// TIA Portal project "OpenLibraryExample" (V13)

(* hardware
DEVICE "S71500/ET200MP station_1"  S7-1500 station
   slot 0: "Rail_0"  6ES7 590-1***0-0AA0
   slot 1: "WaterTreatmentPLC"  CPU 1516-3 PN/DP  6ES7 516-3AN01-0AB0  V1.8
   slot 2: "DI 16x24VDC BA_1"  DI 16x24VDC BA  6ES7 521-1BH10-0AA0  V1.0
   slot 3: "DQ 16x24VDC/0.5A BA_1"  DQ 16x24VDC/0.5A BA  6ES7 522-1BH10-0AA0  V1.0
   slot 4: "AI 4xU/I/RTD/TC ST_1"  AI 4xU/I/RTD/TC ST  6ES7 531-7QD00-0AB0  V1.0
   slot 5: "AQ 4xU/I ST_1"  AQ 4xU/I ST  6ES7 532-5HD00-0AB0  V2.0
DEVICE "SINAMICS G_1"  Sinamics.Device
   slot 0: "	_0"  Rail
   slot 0: "WaterPump"  G120 CU240E-2 PN  6SL3244-0BB12-1FA0  4.7.3
   slot 3: "PM240 IP20"  PM240 IP20  6SL3224-0BE31-5UA0  -
DEVICE "WaterTreatmentHMI"  TP900 Comfort
   slot 0: "HMI"  HMI  6AV2 124-0JC01-0AX0  13.0.1.0
   slot 1: "HMI_RT_1"  TP900 Comfort  6AV2 124-0JC01-0AX0  13.0.1.0
   slot 5: "WaterTreatmentHMI.IE_CP_1"  PROFINET Interface
      slot 1: "PROFINET Interface_1"  PROFINET Interface
         slot 1: "Port_1"  Port
         slot 2: "Port_2"  Port
   slot 7: "WaterTreatmentHMI.MPI/DP_CP_1"  MPI/DP Interface
*)

// ===== PLC "WaterTreatmentPLC"  CPU 1516-3 PN/DP =====

VAR_GLOBAL   // PLC tag table "Open Library"
   "System_Byte" AT %MB1 : Byte;
   "Clock_Byte" AT %MB0 : Byte;
   "Clock_10Hz" AT %M0.0 : Bool;
   "Clock_5Hz" AT %M0.1 : Bool;
   "Clock_2.5Hz" AT %M0.2 : Bool;
   "Clock_2Hz" AT %M0.3 : Bool;
   "Clock_1.25Hz" AT %M0.4 : Bool;
   "Clock_1Hz" AT %M0.5 : Bool;
   "Clock_0.625Hz" AT %M0.6 : Bool;
   "Clock_0.5Hz" AT %M0.7 : Bool;
   "AlwaysTRUE" AT %M1.2 : Bool;
   "AlwaysFALSE" AT %M1.3 : Bool;
   "FirstScan" AT %M1.0 : Bool;
   "DiagStatusUpdate" AT %M1.1 : Bool;
END_VAR

VAR_GLOBAL CONSTANT   // PLC tag table "Open Library"
   "Modes.Auto" : Int := 1;
   "Modes.Manual" : Int := 2;
   "Modes.Independent" : Int := 10;
   "Modes.Stop" : Int := 0;
   "HMI.Status.Stopped" : Int := 0;
   "HMI.Status.Estop" : Int := 1;
   "HMI.Status.Error" : Int := 2;
   "HMI.Status.ForwardWork" : Int := 3;
   "HMI.Status.ReverseHome" : Int := 4;
   "HMI.Status.OnForwardWork" : Int := 5;
   "HMI.Status.OnReverseHome" : Int := 6;
   "IoScaling.S7Analog.Default.iRawMax" : Int := 27648;
   "IoScaling.S7Analog.Default.iRawMin" : Int := 0;
   "IoScaling.S7Analog.Default.bSwapBytes" : Bool := false;
   "IoScaling.S7Analog.+-V/mA.iRawMax" : Int := 27648;
   "IoScaling.S7Analog.+-V/mA.iRawMin" : Int := -27648;
   "IoScaling.S7Analog.Types.Default" : Int := 0;
   "IoScaling.S7Analog.Pt100.iRawMax" : Int := 8500;
   "IoScaling.S7Analog.Pt100.iRawMin" : Int := -2000;
   "IoScaling.S7Analog.Pt100.Climate.iRawMax" : Int := 13000;
   "IoScaling.S7Analog.Pt100.Climate.iRawMin" : Int := -12000;
   "IoScaling.S7Analog.Ni100.iRawMax" : Int := 2500;
   "IoScaling.S7Analog.Ni100.iRawMin" : Int := -600;
   "IoScaling.S7Analog.Ni100.Climate.iRawMax" : Int := 25000;
   "IoScaling.S7Analog.Ni100.Climate.iRawMin" : Int := -6000;
   "IoScaling.S7Analog.Types.+-V/mA" : Int := 1;
   "IoScaling.S7Analog.Types.Pt100" : Int := 2;
   "IoScaling.S7Analog.Types.Pt100.Climate" : Int := 3;
   "IoScaling.S7Analog.Types.Ni100" : Int := 4;
   "IoScaling.S7Analog.Types.Ni100.Climate" : Int := 5;
   "IoScaling.S7Analog.Pt100.rScaledMax" : Real := 850.0;
   "IoScaling.S7Analog.Pt100.rScaledMin" : Real := -200.0;
   "IoScaling.S7Analog.Pt100.Climate.rScaledMax" : Real := 130.0;
   "IoScaling.S7Analog.Pt100.Climate.rScaledMin" : Real := -120.0;
   "IoScaling.S7Analog.Ni100.rScaledMax" : Real := 250.0;
   "IoScaling.S7Analog.Ni100.rScaledMin" : Real := -60.0;
   "IoScaling.S7Analog.Ni100.Climate.rScaledMax" : Real := 250.0;
   "IoScaling.S7Analog.Ni100.Climate.rScaledMin" : Real := -60.0;
   "IoScaling.S7Analog.150Ohms.rScaledMax" : Real := 150.0;
   "IoScaling.S7Analog.150Ohms.rScaledMin" : Real := 0.0;
   "IoScaling.S7Analog.300Ohms.rScaledMax" : Real := 300.0;
   "IoScaling.S7Analog.300Ohms.rScaledMin" : Real := 0.0;
   "IoScaling.S7Analog.600Ohms.rScaledMax" : Real := 600.0;
   "IoScaling.S7Analog.600Ohms.rScaledMin" : Real := 0.0;
   "Estop.MinSetPoint" : Int := 0;
   "Estop.MaxSetPoint" : Int := 1;
   "Estop.HMISetPoint" : Int := 2;
   "Modes.PID.Inactive" : Int := 0;
   "Modes.PID.Pretuning" : Int := 1;
   "Modes.PID.FineTuning" : Int := 2;
   "Modes.PID.AutoMode" : Int := 3;
   "Modes.PID.ManualMode" : Int := 4;
   "HMI.Status.Generic1" : Int := 101;
   "HMI.Status.Generic2" : Int := 102;
   "HMI.Status.Generic3" : Int := 103;
   "HMI.Status.Generic4" : Int := 104;
   "HMI.Status.Generic5" : Int := 105;
   "HMI.Status.GenericNone" : Int := 100;
   "HMI.Status.Generic6" : Int := 106;
   "DataTypes.rMaxReal" : Real := 3.402823e38;
   "DataTypes.rMinReal" : Real := -3.402823e38;
   "DataTypes.iMaxInt" : Int := 32767;
   "DataTypes.iMinInt" : Int := -32768;
END_VAR

VAR_GLOBAL   // PLC tag table "IO"
   "I_MainWaterValveOpen" AT %I0.1 : Bool;   // Main Water Valve Open Feedback
   "I_MainWaterValveClosed" AT %I0.0 : Bool;   // Main Water Valve Closed Feedback
   "Q_MainWaterValveSolenoid" AT %Q0.0 : Bool;   // Main Water Valve Output Solenoid
   "I_WaterPumpContactorAux" AT %I1.0 : Bool;   // Water Pump Contactor Feedback
   "Q_WaterPumpContactor" AT %Q1.0 : Bool;   // Water Pump Contactor Coil
   "I_WaterPumpMSP" AT %I1.1 : Bool;   // Water Pump Motor Protector Feedback
   "I_WaterPumpDisconnect" AT %I1.2 : Bool;   // Water Pump Disconnect Feedback
   "I_WaterPumpCoolingFan" AT %I1.3 : Bool;   // Water Pump Cooling Fan Feedback
   "IW_WaterTemperature" AT %IW50 : Word;   // Water Temperature Actual
   "I_ReturnWaterPumpAux" AT %I0.2 : Bool;   // Return Water Pump Contactor Feedback
   "Q_ReturnWaterPumpContactor" AT %Q0.1 : Bool;   // Return Water Pump Contactor Coil
   "QW_SteamValve" AT %QW50 : Int;   // Water Temperature Steam Analog Valve
   "IW_MainWaterPumpPressure" AT %IW52 : Word;   // Main Water Pump Pressure
   "QW_CoolingCoil" AT %QW52 : Int;   // Water Temperature Cooling Coil
   "QW_RecirculationFan" AT %QW54 : Int;   // Air Recirculation Fan
END_VAR

TYPE "udtOUT_PIDInterface"
   STRUCT
      rProcessValue : Real;
      wProcessValue : Word;
      rSetPoint : Real;
      rManualValue : Real;
      iModeRequest : Int;
      bManualEnable : Bool;
      bModeChangeRequest : Bool;
   END_STRUCT;
END_TYPE

// folder: Error

TYPE "udtError_AnalogInput"
   STRUCT
      LowLowAlarm : Bool;
      HighHighAlarm : Bool;
      Invalid : Bool;
   END_STRUCT;
END_TYPE

TYPE "udtError_AnalogOutput"
   STRUCT
      OutOfRange : Bool;
      ConfigurationError : Bool;
   END_STRUCT;
END_TYPE

TYPE "udtError_Motor"
   STRUCT
      MotorProtectorTripped : Bool;
      LocalDisconnectOff : Bool;
      ClutchTripped : Bool;
      NoSignalForward : Bool;
      NoSignalReverse : Bool;
      MotorNotStopped : Bool;
   END_STRUCT;
END_TYPE

TYPE "udtError_AnalogValve"
   STRUCT
      InvalidFeedback : Bool;
   END_STRUCT;
END_TYPE

TYPE "udtError_Valve"
   STRUCT
      NoHomeFeedback : Bool;
      NoWorkFeedback : Bool;
      HomeFeedbackStillActive : Bool;
      WorkFeedbackStillActive : Bool;
   END_STRUCT;
END_TYPE

TYPE "udtError_VFD"
   STRUCT
      MotorProtectorTripped : Bool;
      LocalDisconnectOff : Bool;
      ClutchTripped : Bool;
      NoContactorFeedback : Bool;
      ContactorStillOn : Bool;
      NoSignalForward : Bool;
      NoSignalReverse : Bool;
      MotorNotStopped : Bool;
      MaxFrequencyReached : Bool;
      Overcurrent : Bool;
      MotorOverload : Bool;
      VFDOverload : Bool;
      GeneralFault : Bool;
      NoCoolingFanFeedback : Bool;
   END_STRUCT;
END_TYPE

TYPE "udtError_PID"
   STRUCT
      InputOutOfRange : Bool;
      InputPERInvalid : Bool;
      ValueOscillationFailed : Bool;
      ProcessValueCloseToSetPoint : Bool;
      SetPointChangedDuringTuning : Bool;
      PretuningDuringFineTuning : Bool;
      InvalidOutputValueLimits : Bool;
      InvalidFineTuningParameter : Bool;
      InputInvalidFormat : Bool;
      OutputCalculationError : Bool;
      SamplingTimeError : Bool;
      SetPointInvalidFormat : Bool;
      ManualInvalidFormat : Bool;
      SubstituteOutputInvalidFormat : Bool;
      DisturbanceInvalidFormat : Bool;
   END_STRUCT;
END_TYPE

// folder: HMI

TYPE "udtHMI_VFD_Control"
   STRUCT
      iMode : Int;
      iErrorCode : Int;
      iStatus : Int;
      rManualSpeedSP : Real;
      rAutoSpeedSP : Real;
      rActualSpeed : Real;
      rActualCurrent : Real;
      rActualPower : Real;
      bPB_ResetError : Bool;
      bPB_Forward : Bool;
      bPB_Reverse : Bool;
      bPB_Stop : Bool;
      bPBEN_ResetError : Bool;
      bPBEN_Forward : Bool;
      bPBEN_Reverse : Bool;
      bPBEN_Stop : Bool;
      bForwardOn : Bool;
      bReverseOn : Bool;
      bSignalForward : Bool;
      bSignalReverse : Bool;
      bError : Bool;
      bInterlock : Bool;
   END_STRUCT;
END_TYPE

TYPE "udtHMI_AnalogInput"
   STRUCT
      iMode : Int;
      iErrorCode : Int;
      iStatus : Int;
      rActiveValue : Real;
      rInputValue : Real;
      rManualValue : Real;
      bPB_ResetError : Bool;
      bPBEN_ResetError : Bool;
      bError : Bool;
   END_STRUCT;
END_TYPE

TYPE "udtHMI_MotorControl"
   STRUCT
      iMode : Int;
      iErrorCode : Int;
      iStatus : Int;
      bPB_ResetError : Bool;
      bPB_Forward : Bool;
      bPB_Reverse : Bool;
      bPB_Stop : Bool;
      bPBEN_ResetError : Bool;
      bPBEN_Forward : Bool;
      bPBEN_Reverse : Bool;
      bPBEN_Stop : Bool;
      bForwardOn : Bool;
      bReverseOn : Bool;
      bSignalForward : Bool;
      bSignalReverse : Bool;
      bError : Bool;
      bInterlock : Bool;
   END_STRUCT;
END_TYPE

TYPE "udtHMI_ValveControl"
   STRUCT
      iMode : Int;
      iErrorCode : Int;
      iStatus : Int;
      bPB_ResetError : Bool;
      bPB_Home : Bool;
      bPB_Work : Bool;
      bPBEN_ResetError : Bool;
      bPBEN_Home : Bool;
      bPBEN_Work : Bool;
      bHomeOn : Bool;
      bWorkOn : Bool;
      bSignalHome : Bool;
      bSignalWork : Bool;
      bError : Bool;
      bInterlock : Bool;
   END_STRUCT;
END_TYPE

TYPE "udtHMI_PIDControlParameters"
   STRUCT
      rProportionalGain : Real;
      rIntegralTime : Real;
      rDerivativeTime : Real;
      rProportionalWeight : Real;
      rDerivativeWeight : Real;
   END_STRUCT;
END_TYPE

TYPE "udtHMI_Interlock"
   STRUCT
      abInterlocks : Array[1..16] of Bool;
      asInterlockNames : Array[1..16] of String[20];
      bInterlockOk : Bool;
   END_STRUCT;
END_TYPE

TYPE "udtHMI_SystemControl"
VERSION : 0.1
   STRUCT
      iMode : Int;
      bEStop : Bool;
      bError : Bool;
      bAuto : Bool;
      bIndependentEnable : Bool;
      bPB_ResetError : Bool;
   END_STRUCT;
END_TYPE

TYPE "udtHMI_PIDInterface"
   STRUCT
      iMode : Int;
      iPIDMode : Int;
      iErrorCode : Int;
      iEstopFunction : Int;
      rEstopValue : Real;
      rManualSP : Real;
      rAutoSP : Real;
      rActualInput : Real;
      wActualInputPeripheral : Word;
      rOutput : Real;
      wOutputPeripheral : Word;
      bPB_ResetError : Bool;
      bPB_Pretune : Bool;
      bPB_FineTune : Bool;
      bPB_AutomaticMode : Bool;
      bPB_ManualMode : Bool;
      bPB_ManualTuning : Bool;
      bTOG_ManualTuning : Bool;
      bPBEN_ResetError : Bool;
      bPBEN_Pretune : Bool;
      bPBEN_FineTune : Bool;
      bPBEN_AutomaticMode : Bool;
      bPBEN_ManualMode : Bool;
      bError : Bool;
      bErrorAck : Bool;
      PID_ControlParameters : "udtHMI_PIDControlParameters";
   END_STRUCT;
END_TYPE

TYPE "udtHMI_AnalogOutput"
   STRUCT
      iMode : Int;
      iErrorCode : Int;
      rValue : Real;
      rAutoValue : Real;
      rManualValue : Real;
      rEstopValue : Real;
      bPB_ResetError : Bool;
      bPBEN_ResetError : Bool;
      bError : Bool;
      bInterlock : Bool;
      iEstopFunction : Int;
   END_STRUCT;
END_TYPE

TYPE "udtHMI_AnalogValveControl"
   STRUCT
      iMode : Int;
      iErrorCode : Int;
      iStatus : Int;
      rManualSP : Real;
      rAutoSP : Real;
      rEstopSP : Real;
      rActual : Real;
      bPB_ResetError : Bool;
      bPBEN_ResetError : Bool;
      bError : Bool;
      bInterlock : Bool;
      iEstopFunction : Int;
   END_STRUCT;
END_TYPE

// folder: Systems/Data

DATA_BLOCK "dbWaterSystem"   // DB610
{ S7_Optimized_Access := 'FALSE' }
VERSION : 0.1
   VAR
      SOL_MainWater : "udtHMI_ValveControl";
      VFD_WaterPump : "udtHMI_VFD_Control";
      INT_WaterPump : "udtHMI_Interlock";
      AI_WaterPumpPressure : "udtHMI_AnalogInput";
      MTR_ReturnWaterPump : "udtHMI_MotorControl";
      ANA_SteamValve : "udtHMI_AnalogValveControl";
      AO_CoolingCoil : "udtHMI_AnalogOutput";
      SystemControl : "udtHMI_SystemControl";
      WaterTemperature : Struct
      END_STRUCT;
   END_VAR
BEGIN
END_DATA_BLOCK

DATA_BLOCK "dbAirSystem"   // DB620
{ S7_Optimized_Access := 'FALSE' }
VERSION : 0.1
   VAR
      SystemControl : "udtHMI_SystemControl";
      VFD_RecirculationFan : "udtHMI_VFD_Control";
   END_VAR
BEGIN
END_DATA_BLOCK

DATA_BLOCK "dbErrors_WaterSystem"   // DB710
{ S7_Optimized_Access := 'FALSE' }
VERSION : 0.1
   VAR
      SOL_MainWater : "udtError_Valve";
      VFD_WaterPump : "udtError_VFD";
      AI_WaterPumpPressure : "udtError_AnalogInput";
      MTR_ReturnWaterPump : "udtError_Motor";
      ANA_SteamValve : "udtError_AnalogValve";
      AO_CoolingCoil : "udtError_AnalogOutput";
      PID_WaterTemperature : "udtError_PID";
      AI_WaterTemperature : "udtError_AnalogInput";
      bMainPumpHighHighPressure : Bool;
      bMainPumpHighPressure : Bool;
   END_VAR
BEGIN
END_DATA_BLOCK

DATA_BLOCK "dbErrors_AirSystem"   // DB720
{ S7_Optimized_Access := 'FALSE' }
VERSION : 0.1
   VAR
      VFD_RecirculationFan : "udtError_VFD";
   END_VAR
BEGIN
END_DATA_BLOCK

// folder: Systems/Instance Data

DATA_BLOCK "dbIns_Master"   // DB1
{ S7_Optimized_Access := 'FALSE' }
VERSION : 0.1
// stored: InstanceOfName fbMaster
"fbMaster"
BEGIN
END_DATA_BLOCK

DATA_BLOCK "dbIns_CyclicInterrupt"   // DB30
{ S7_Optimized_Access := 'FALSE' }
VERSION : 0.1
// stored: InstanceOfName fbCyclicInterrupt
"fbCyclicInterrupt"
BEGIN
END_DATA_BLOCK

DATA_BLOCK "dbIns_WaterSystem"   // DB510
{ S7_Optimized_Access := 'FALSE' }
VERSION : 0.1
// stored: InstanceOfName fbWaterSystem
"fbWaterSystem"
BEGIN
END_DATA_BLOCK

DATA_BLOCK "dbIns_AirSystem"   // DB520
{ S7_Optimized_Access := 'FALSE' }
VERSION : 0.1
// stored: InstanceOfName fbAirSystem
"fbAirSystem"
BEGIN
END_DATA_BLOCK

// folder: Library Blocks/Devices

FUNCTION_BLOCK "fbValve_Solenoid"   // FB110, LAD
TITLE = Controls a double- or single-acting valve
{ S7_Optimized_Access := 'FALSE' }
VERSION : 0.1
   VAR_TEMP   // added for the SCL form of the ladder/FBD networks
      _w1 : Bool;
      _w2 : Bool;
   END_VAR
BEGIN

REGION Network 1: --------------------------------------------------------- Inputs ------------------------------------------------------------------
END_REGION

REGION Network 2: Read HMI input buttons
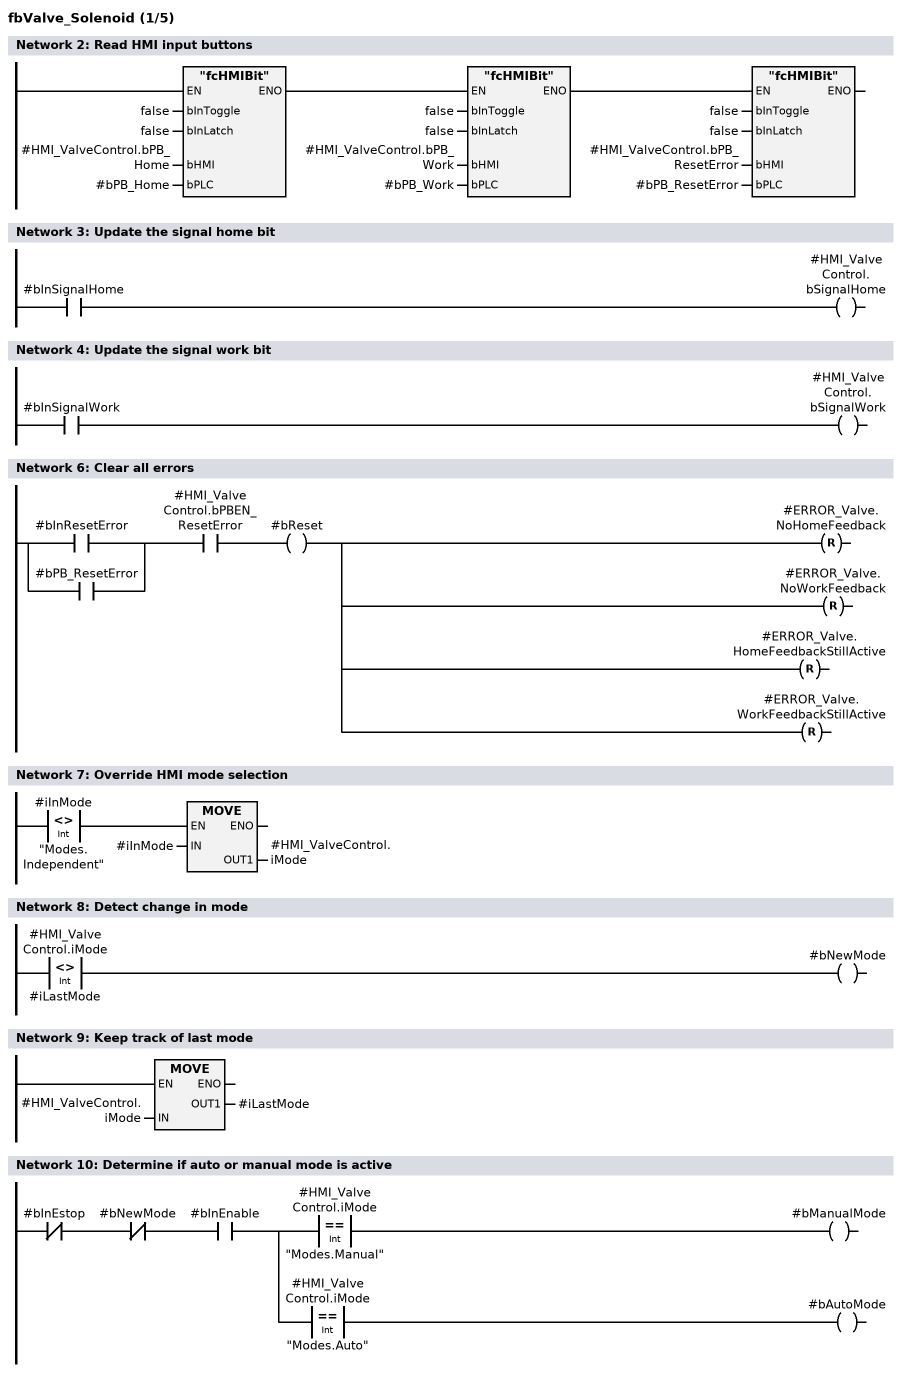
   RUNG wire#powerrail
      "fcHMIBit"(bInToggle := false, bInLatch := false, bHMI := #HMI_ValveControl.bPB_Home, bPLC := #bPB_Home)
      "fcHMIBit"(bInToggle := false, bInLatch := false, bHMI := #HMI_ValveControl.bPB_Work, bPLC := #bPB_Work)
      "fcHMIBit"(bInToggle := false, bInLatch := false, bHMI := #HMI_ValveControl.bPB_ResetError, bPLC := #bPB_ResetError)
   END_RUNG
   // the same network as SCL:
   "fcHMIBit"(bInToggle := false,
              bInLatch := false,
              bHMI := #HMI_ValveControl.bPB_Home,
              bPLC := #bPB_Home,
              ENO => #_w1);
   "fcHMIBit"(EN := #_w1,
              bInToggle := false,
              bInLatch := false,
              bHMI := #HMI_ValveControl.bPB_Work,
              bPLC := #bPB_Work,
              ENO => #_w2);
   IF #_w2 THEN
       "fcHMIBit"(bInToggle := false,
                  bInLatch := false,
                  bHMI := #HMI_ValveControl.bPB_ResetError,
                  bPLC := #bPB_ResetError);
   END_IF;
END_REGION

REGION Network 3: Update the signal home bit
   RUNG wire#powerrail
      Contact( #bInSignalHome )
      Coil( #HMI_ValveControl.bSignalHome )
   END_RUNG
   // the same network as SCL:
   #HMI_ValveControl.bSignalHome := #bInSignalHome;
END_REGION

REGION Network 4: Update the signal work bit
   RUNG wire#powerrail
      Contact( #bInSignalWork )
      Coil( #HMI_ValveControl.bSignalWork )
   END_RUNG
   // the same network as SCL:
   #HMI_ValveControl.bSignalWork := #bInSignalWork;
END_REGION

REGION Network 5: --------------------------------------------------- Control Logic ------------------------------------------------------------
END_REGION

REGION Network 6: Clear all errors
   RUNG wire#powerrail
      Contact( #bInResetError )
      wire#w1
      Contact( #HMI_ValveControl.bPBEN_ResetError )
      Coil( #bReset )
      wire#w2
      R_Coil( #ERROR_Valve.NoHomeFeedback )
   END_RUNG
   RUNG wire#powerrail
      Contact( #bPB_ResetError )
   END_RUNG wire#w1
   RUNG wire#w2
      R_Coil( #ERROR_Valve.NoWorkFeedback )
   END_RUNG
   RUNG wire#w2
      R_Coil( #ERROR_Valve.HomeFeedbackStillActive )
   END_RUNG
   RUNG wire#w2
      R_Coil( #ERROR_Valve.WorkFeedbackStillActive )
   END_RUNG
   // the same network as SCL:
   #bReset := (#bInResetError OR #bPB_ResetError) AND #HMI_ValveControl.bPBEN_ResetError;
   IF #bReset THEN
       #ERROR_Valve.NoHomeFeedback := FALSE;
       #ERROR_Valve.NoWorkFeedback := FALSE;
       #ERROR_Valve.HomeFeedbackStillActive := FALSE;
       #ERROR_Valve.WorkFeedbackStillActive := FALSE;
   END_IF;
END_REGION

REGION Network 7: Override HMI mode selection
   RUNG wire#powerrail
      { S7_Templates := "SrcType := Int" } NE_Contact(in1 := #iInMode, in2 := "Modes.Independent")
      { S7_GenerateENO := "TRUE" } Move(in := #iInMode, out1 => #HMI_ValveControl.iMode)
   END_RUNG
   // the same network as SCL:
   IF #iInMode <> "Modes.Independent" THEN #HMI_ValveControl.iMode := #iInMode; END_IF;
END_REGION

REGION Network 8: Detect change in mode
   RUNG wire#powerrail
      { S7_Templates := "SrcType := Int" } NE_Contact(in1 := #HMI_ValveControl.iMode, in2 := #iLastMode)
      Coil( #bNewMode )
   END_RUNG
   // the same network as SCL:
   #bNewMode := #HMI_ValveControl.iMode <> #iLastMode;
END_REGION

REGION Network 9: Keep track of last mode
   RUNG wire#powerrail
      { S7_GenerateENO := "TRUE" } Move(in := #HMI_ValveControl.iMode, out1 => #iLastMode)
   END_RUNG
   // the same network as SCL:
   #iLastMode := #HMI_ValveControl.iMode;
END_REGION

REGION Network 10: Determine if auto or manual mode is active
   RUNG wire#powerrail
      I_Contact( #bInEstop )
      I_Contact( #bNewMode )
      Contact( #bInEnable )
      wire#w1
      { S7_Templates := "SrcType := Int" } EQ_Contact(in1 := #HMI_ValveControl.iMode, in2 := "Modes.Manual")
      Coil( #bManualMode )
   END_RUNG
   RUNG wire#w1
      { S7_Templates := "SrcType := Int" } EQ_Contact(in1 := #HMI_ValveControl.iMode, in2 := "Modes.Auto")
      Coil( #bAutoMode )
   END_RUNG
   // the same network as SCL:
   #_w1 := NOT #bInEstop AND NOT #bNewMode AND #bInEnable;
   #bManualMode := #_w1 AND (#HMI_ValveControl.iMode = "Modes.Manual");
   #bAutoMode := #_w1 AND (#HMI_ValveControl.iMode = "Modes.Auto");
END_REGION

REGION Network 11: Enable Home & Work Positions
   // IF manual mode AND no estop AND not a new mode AND enabled => 
   // --if no cylinder errors, enable move to Home and Work
   // --enable home and work HMI buttons only in manual mode
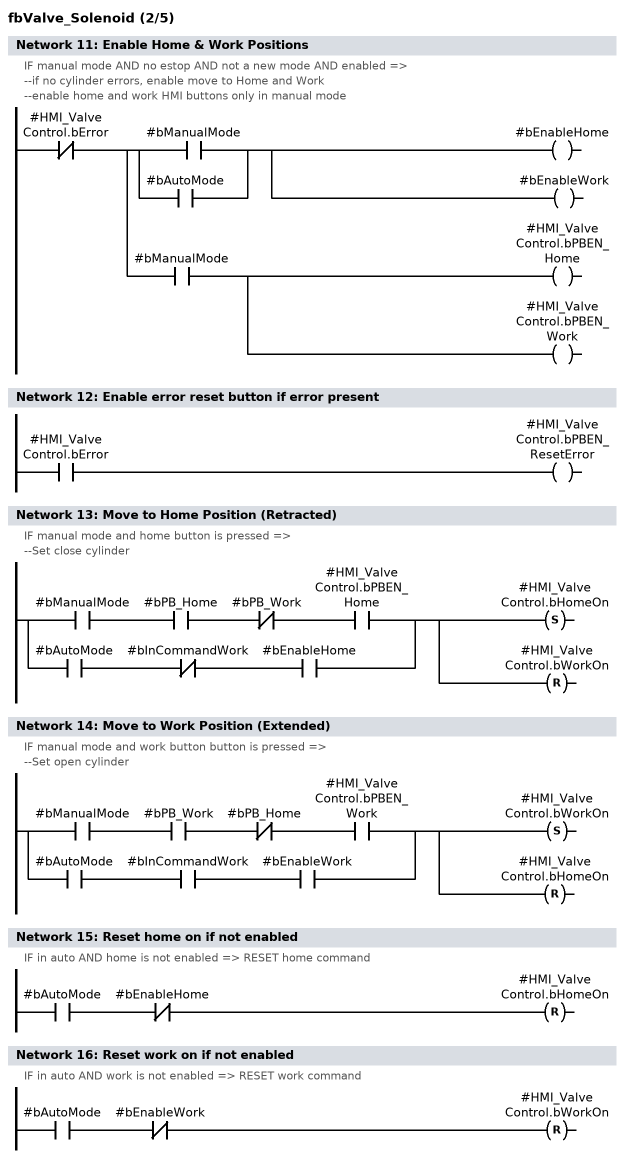
   RUNG wire#powerrail
      I_Contact( #HMI_ValveControl.bError )
      wire#w1
      Contact( #bManualMode )
      wire#w2
      Coil( #bEnableHome )
   END_RUNG
   RUNG wire#w1
      Contact( #bAutoMode )
   END_RUNG wire#w2
   RUNG wire#w2
      Coil( #bEnableWork )
   END_RUNG
   RUNG wire#w1
      Contact( #bManualMode )
      wire#w3
      Coil( #HMI_ValveControl.bPBEN_Home )
   END_RUNG
   RUNG wire#w3
      Coil( #HMI_ValveControl.bPBEN_Work )
   END_RUNG
   // the same network as SCL:
   #_w1 := NOT #HMI_ValveControl.bError;
   #bEnableHome := #_w1 AND (#bManualMode OR #bAutoMode);
   #bEnableWork := #bEnableHome;
   #HMI_ValveControl.bPBEN_Home := #_w1 AND #bManualMode;
   #HMI_ValveControl.bPBEN_Work := #HMI_ValveControl.bPBEN_Home;
END_REGION

REGION Network 12: Enable error reset button if error present
   RUNG wire#powerrail
      Contact( #HMI_ValveControl.bError )
      Coil( #HMI_ValveControl.bPBEN_ResetError )
   END_RUNG
   // the same network as SCL:
   #HMI_ValveControl.bPBEN_ResetError := #HMI_ValveControl.bError;
END_REGION

REGION Network 13: Move to Home Position (Retracted)
   // IF manual mode and home button is pressed =>
   // --Set close cylinder
   RUNG wire#powerrail
      Contact( #bManualMode )
      Contact( #bPB_Home )
      I_Contact( #bPB_Work )
      Contact( #HMI_ValveControl.bPBEN_Home )
      wire#w1
      S_Coil( #HMI_ValveControl.bHomeOn )
   END_RUNG
   RUNG wire#powerrail
      Contact( #bAutoMode )
      I_Contact( #bInCommandWork )
      Contact( #bEnableHome )
   END_RUNG wire#w1
   RUNG wire#w1
      R_Coil( #HMI_ValveControl.bWorkOn )
   END_RUNG
   // the same network as SCL:
   IF (#bManualMode AND #bPB_Home AND NOT #bPB_Work AND #HMI_ValveControl.bPBEN_Home) OR (#bAutoMode AND NOT #bInCommandWork AND #bEnableHome) THEN
       #HMI_ValveControl.bHomeOn := TRUE;
       #HMI_ValveControl.bWorkOn := FALSE;
   END_IF;
END_REGION

REGION Network 14: Move to Work Position (Extended)
   // IF manual mode and work button button is pressed =>
   // --Set open cylinder
   RUNG wire#powerrail
      Contact( #bManualMode )
      Contact( #bPB_Work )
      I_Contact( #bPB_Home )
      Contact( #HMI_ValveControl.bPBEN_Work )
      wire#w1
      S_Coil( #HMI_ValveControl.bWorkOn )
   END_RUNG
   RUNG wire#powerrail
      Contact( #bAutoMode )
      Contact( #bInCommandWork )
      Contact( #bEnableWork )
   END_RUNG wire#w1
   RUNG wire#w1
      R_Coil( #HMI_ValveControl.bHomeOn )
   END_RUNG
   // the same network as SCL:
   IF (#bManualMode AND #bPB_Work AND NOT #bPB_Home AND #HMI_ValveControl.bPBEN_Work) OR (#bAutoMode AND #bInCommandWork AND #bEnableWork) THEN
       #HMI_ValveControl.bWorkOn := TRUE;
       #HMI_ValveControl.bHomeOn := FALSE;
   END_IF;
END_REGION

REGION Network 15: Reset home on if not enabled
   // IF in auto AND home is not enabled => RESET home command
   RUNG wire#powerrail
      Contact( #bAutoMode )
      I_Contact( #bEnableHome )
      R_Coil( #HMI_ValveControl.bHomeOn )
   END_RUNG
   // the same network as SCL:
   IF #bAutoMode AND NOT #bEnableHome THEN #HMI_ValveControl.bHomeOn := FALSE; END_IF;
END_REGION

REGION Network 16: Reset work on if not enabled
   // IF in auto AND work is not enabled => RESET work command
   RUNG wire#powerrail
      Contact( #bAutoMode )
      I_Contact( #bEnableWork )
      R_Coil( #HMI_ValveControl.bWorkOn )
   END_RUNG
   // the same network as SCL:
   IF #bAutoMode AND NOT #bEnableWork THEN #HMI_ValveControl.bWorkOn := FALSE; END_IF;
END_REGION

REGION Network 17: Reset both home and work if not in auto or manual
   // IF not in auto AND not in manual => RESET home and work commands
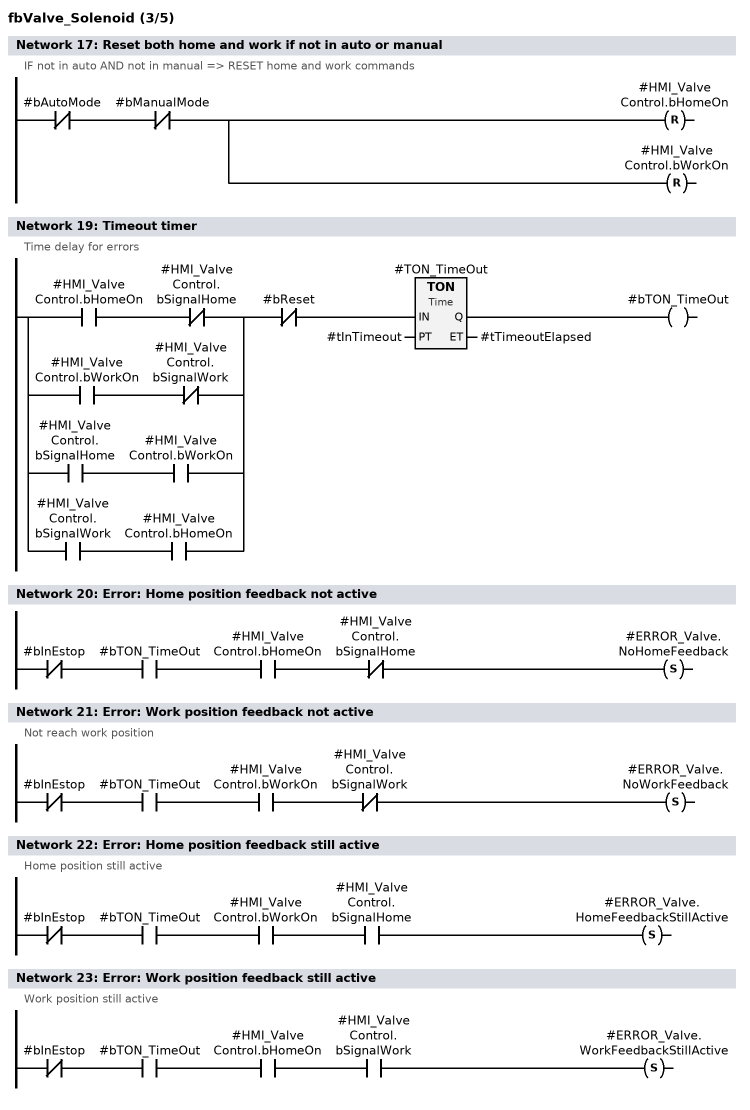
   RUNG wire#powerrail
      I_Contact( #bAutoMode )
      I_Contact( #bManualMode )
      wire#w1
      R_Coil( #HMI_ValveControl.bHomeOn )
   END_RUNG
   RUNG wire#w1
      R_Coil( #HMI_ValveControl.bWorkOn )
   END_RUNG
   // the same network as SCL:
   IF NOT #bAutoMode AND NOT #bManualMode THEN
       #HMI_ValveControl.bHomeOn := FALSE;
       #HMI_ValveControl.bWorkOn := FALSE;
   END_IF;
END_REGION

REGION Network 18: --------------------------------------------------------- Errors ------------------------------------------------------------------
END_REGION

REGION Network 19: Timeout timer
   // Time delay for errors
   #TON_TimeOut.TON(IN := ((#HMI_ValveControl.bHomeOn AND NOT #HMI_ValveControl.bSignalHome) OR (#HMI_ValveControl.bWorkOn AND NOT #HMI_ValveControl.bSignalWork) OR (#HMI_ValveControl.bSignalHome AND #HMI_ValveControl.bWorkOn) OR (#HMI_ValveControl.bSignalWork AND #HMI_ValveControl.bHomeOn)) AND NOT #bReset,
                    PT := #tInTimeout,
                    ET => #tTimeoutElapsed);
   #bTON_TimeOut := #TON_TimeOut.Q;
END_REGION

REGION Network 20: Error: Home position feedback not active
   RUNG wire#powerrail
      I_Contact( #bInEstop )
      Contact( #bTON_TimeOut )
      Contact( #HMI_ValveControl.bHomeOn )
      I_Contact( #HMI_ValveControl.bSignalHome )
      S_Coil( #ERROR_Valve.NoHomeFeedback )
   END_RUNG
   // the same network as SCL:
   IF NOT #bInEstop AND #bTON_TimeOut AND #HMI_ValveControl.bHomeOn AND NOT #HMI_ValveControl.bSignalHome THEN
       #ERROR_Valve.NoHomeFeedback := TRUE;
   END_IF;
END_REGION

REGION Network 21: Error: Work position feedback not active
   // Not reach work position
   RUNG wire#powerrail
      I_Contact( #bInEstop )
      Contact( #bTON_TimeOut )
      Contact( #HMI_ValveControl.bWorkOn )
      I_Contact( #HMI_ValveControl.bSignalWork )
      S_Coil( #ERROR_Valve.NoWorkFeedback )
   END_RUNG
   // the same network as SCL:
   IF NOT #bInEstop AND #bTON_TimeOut AND #HMI_ValveControl.bWorkOn AND NOT #HMI_ValveControl.bSignalWork THEN
       #ERROR_Valve.NoWorkFeedback := TRUE;
   END_IF;
END_REGION

REGION Network 22: Error: Home position feedback still active
   // Home position still active
   RUNG wire#powerrail
      I_Contact( #bInEstop )
      Contact( #bTON_TimeOut )
      Contact( #HMI_ValveControl.bWorkOn )
      Contact( #HMI_ValveControl.bSignalHome )
      S_Coil( #ERROR_Valve.HomeFeedbackStillActive )
   END_RUNG
   // the same network as SCL:
   IF NOT #bInEstop AND #bTON_TimeOut AND #HMI_ValveControl.bWorkOn AND #HMI_ValveControl.bSignalHome THEN
       #ERROR_Valve.HomeFeedbackStillActive := TRUE;
   END_IF;
END_REGION

REGION Network 23: Error: Work position feedback still active
   // Work position still active
   RUNG wire#powerrail
      I_Contact( #bInEstop )
      Contact( #bTON_TimeOut )
      Contact( #HMI_ValveControl.bHomeOn )
      Contact( #HMI_ValveControl.bSignalWork )
      S_Coil( #ERROR_Valve.WorkFeedbackStillActive )
   END_RUNG
   // the same network as SCL:
   IF NOT #bInEstop AND #bTON_TimeOut AND #HMI_ValveControl.bHomeOn AND #HMI_ValveControl.bSignalWork THEN
       #ERROR_Valve.WorkFeedbackStillActive := TRUE;
   END_IF;
END_REGION

REGION Network 24: Error scroller
   // Call the Error-Scroller which cyles through all possible errors and checks 
   // their state for display on the HMI
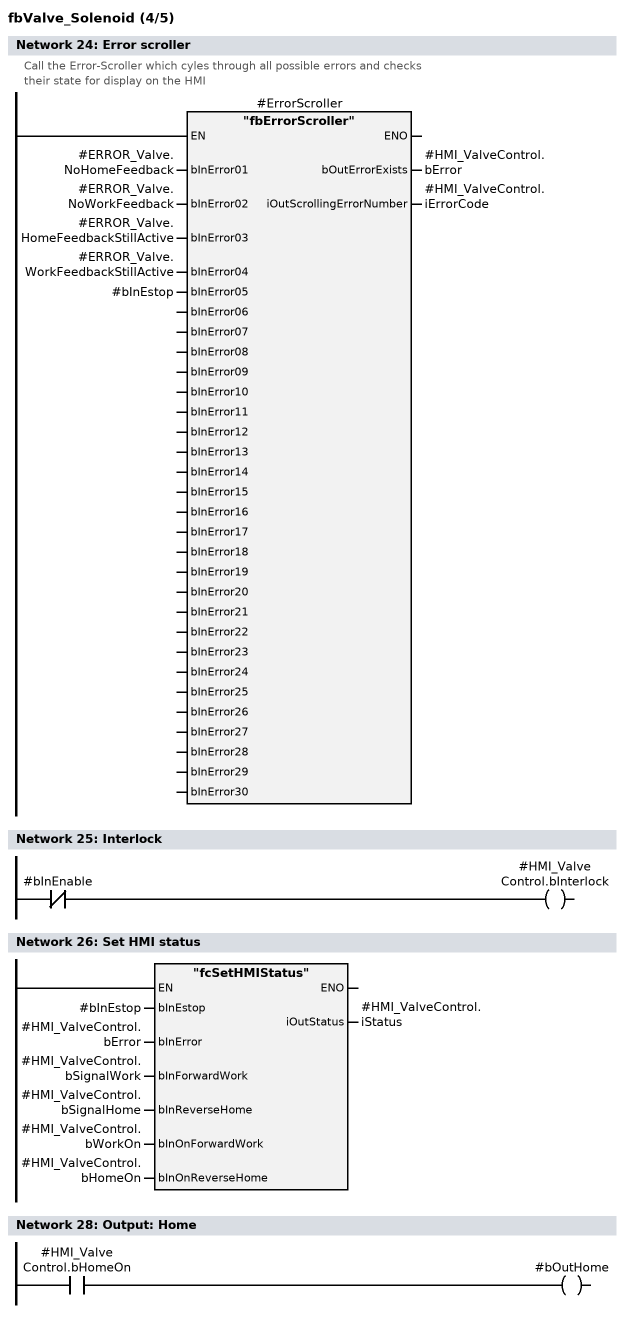
   RUNG wire#powerrail
      #ErrorScroller(bInError01 := #ERROR_Valve.NoHomeFeedback, bInError02 := #ERROR_Valve.NoWorkFeedback, bInError03 := #ERROR_Valve.HomeFeedbackStillActive, bInError04 := #ERROR_Valve.WorkFeedbackStillActive, bInError05 := #bInEstop, bInError06 :=, bInError07 :=, bInError08 :=, bInError09 :=, bInError10 :=, bInError11 :=, bInError12 :=, bInError13 :=, bInError14 :=, bInError15 :=, bInError16 :=, bInError17 :=, bInError18 :=, bInError19 :=, bInError20 :=, bInError21 :=, bInError22 :=, bInError23 :=, bInError24 :=, bInError25 :=, bInError26 :=, bInError27 :=, bInError28 :=, bInError29 :=, bInError30 :=, bOutErrorExists => #HMI_ValveControl.bError, iOutScrollingErrorNumber => #HMI_ValveControl.iErrorCode)
   END_RUNG
   // the same network as SCL:
   #ErrorScroller(bInError01 := #ERROR_Valve.NoHomeFeedback,   // "fbErrorScroller"
                  bInError02 := #ERROR_Valve.NoWorkFeedback,
                  bInError03 := #ERROR_Valve.HomeFeedbackStillActive,
                  bInError04 := #ERROR_Valve.WorkFeedbackStillActive,
                  bInError05 := #bInEstop,
                  bOutErrorExists => #HMI_ValveControl.bError,
                  iOutScrollingErrorNumber => #HMI_ValveControl.iErrorCode);
END_REGION

REGION Network 25: Interlock
   RUNG wire#powerrail
      I_Contact( #bInEnable )
      Coil( #HMI_ValveControl.bInterlock )
   END_RUNG
   // the same network as SCL:
   #HMI_ValveControl.bInterlock := NOT #bInEnable;
END_REGION

REGION Network 26: Set HMI status
   RUNG wire#powerrail
      "fcSetHMIStatus"(bInEstop := #bInEstop, bInError := #HMI_ValveControl.bError, bInForwardWork := #HMI_ValveControl.bSignalWork, bInReverseHome := #HMI_ValveControl.bSignalHome, bInOnForwardWork := #HMI_ValveControl.bWorkOn, bInOnReverseHome := #HMI_ValveControl.bHomeOn, iOutStatus => #HMI_ValveControl.iStatus)
   END_RUNG
   // the same network as SCL:
   "fcSetHMIStatus"(bInEstop := #bInEstop,
                    bInError := #HMI_ValveControl.bError,
                    bInForwardWork := #HMI_ValveControl.bSignalWork,
                    bInReverseHome := #HMI_ValveControl.bSignalHome,
                    bInOnForwardWork := #HMI_ValveControl.bWorkOn,
                    bInOnReverseHome := #HMI_ValveControl.bHomeOn,
                    iOutStatus => #HMI_ValveControl.iStatus);
END_REGION

REGION Network 27: -------------------------------------------------- Outputs --------------------------------------------------
END_REGION

REGION Network 28: Output: Home
   RUNG wire#powerrail
      Contact( #HMI_ValveControl.bHomeOn )
      Coil( #bOutHome )
   END_RUNG
   // the same network as SCL:
   #bOutHome := #HMI_ValveControl.bHomeOn;
END_REGION

REGION Network 29: Output: Work
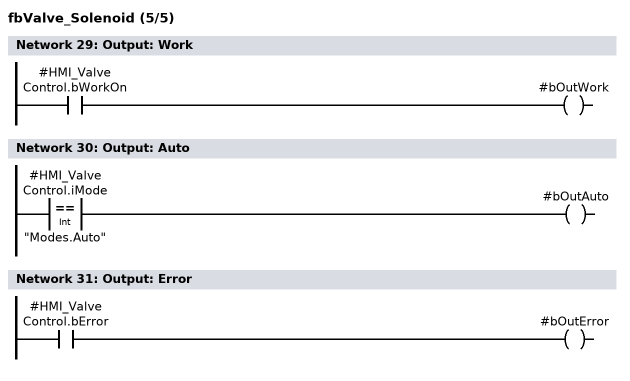
   RUNG wire#powerrail
      Contact( #HMI_ValveControl.bWorkOn )
      Coil( #bOutWork )
   END_RUNG
   // the same network as SCL:
   #bOutWork := #HMI_ValveControl.bWorkOn;
END_REGION

REGION Network 30: Output: Auto
   RUNG wire#powerrail
      { S7_Templates := "SrcType := Int" } EQ_Contact(in1 := #HMI_ValveControl.iMode, in2 := "Modes.Auto")
      Coil( #bOutAuto )
   END_RUNG
   // the same network as SCL:
   #bOutAuto := #HMI_ValveControl.iMode = "Modes.Auto";
END_REGION

REGION Network 31: Output: Error
   RUNG wire#powerrail
      Contact( #HMI_ValveControl.bError )
      Coil( #bOutError )
   END_RUNG
   // the same network as SCL:
   #bOutError := #HMI_ValveControl.bError;
END_REGION
END_FUNCTION_BLOCK

FUNCTION_BLOCK "fbValve_Analog"   // FB111, LAD
TITLE = Controls an analog valve
{ S7_Optimized_Access := 'FALSE' }
VERSION : 0.1
   VAR_TEMP   // added for the SCL form of the ladder/FBD networks
      _w1 : Bool;
      _w2 : Bool;
      _w3 : Bool;
      _w4 : Bool;
   END_VAR
BEGIN

REGION Network 1: Read HMI input buttons
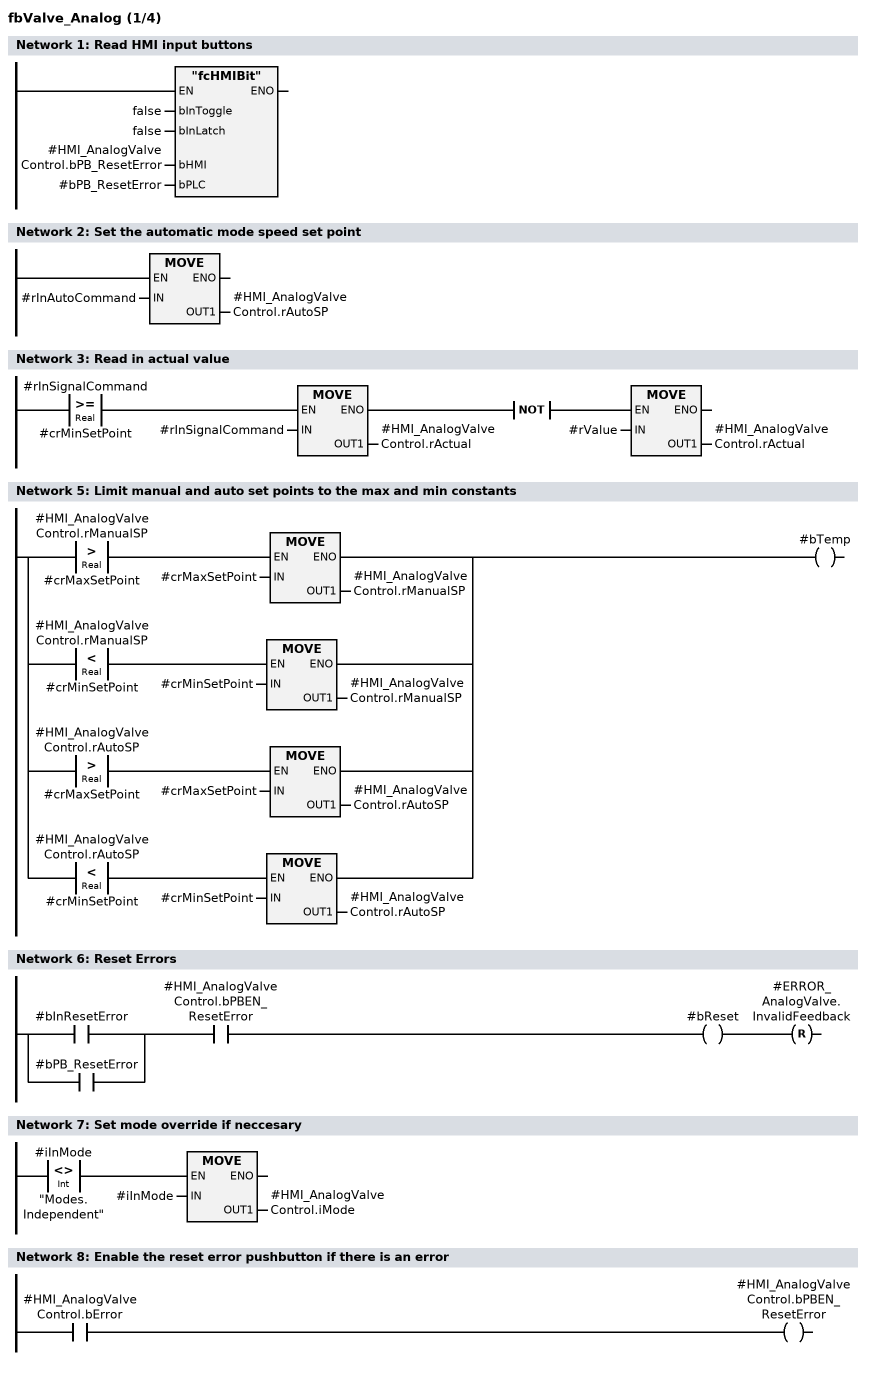
   RUNG wire#powerrail
      "fcHMIBit"(bInToggle := false, bInLatch := false, bHMI := #HMI_AnalogValveControl.bPB_ResetError, bPLC := #bPB_ResetError)
   END_RUNG
   // the same network as SCL:
   "fcHMIBit"(bInToggle := false,
              bInLatch := false,
              bHMI := #HMI_AnalogValveControl.bPB_ResetError,
              bPLC := #bPB_ResetError);
END_REGION

REGION Network 2: Set the automatic mode speed set point
   RUNG wire#powerrail
      { S7_GenerateENO := "TRUE" } Move(in := #rInAutoCommand, out1 => #HMI_AnalogValveControl.rAutoSP)
   END_RUNG
   // the same network as SCL:
   #HMI_AnalogValveControl.rAutoSP := #rInAutoCommand;
END_REGION

REGION Network 3: Read in actual value
   RUNG wire#powerrail
      { S7_Templates := "SrcType := Real" } GE_Contact(in1 := #rInSignalCommand, in2 := #crMinSetPoint)
      { S7_GenerateENO := "TRUE" } Move(in := #rInSignalCommand, out1 => #HMI_AnalogValveControl.rActual)
      Not()
      { S7_GenerateENO := "TRUE" } Move(in := #rValue, out1 => #HMI_AnalogValveControl.rActual)
   END_RUNG
   // the same network as SCL:
   // ENO of a box is taken as its EN; it also drops when the box reports an error
   #_w1 := #rInSignalCommand >= #crMinSetPoint;
   IF #_w1 THEN #HMI_AnalogValveControl.rActual := #rInSignalCommand; END_IF;
   IF NOT #_w1 THEN #HMI_AnalogValveControl.rActual := #rValue; END_IF;
END_REGION

REGION Network 4: --------------------------------------------------- Control Logic ------------------------------------------------------------
END_REGION

REGION Network 5: Limit manual and auto set points to the max and min constants
   RUNG wire#powerrail
      { S7_Templates := "SrcType := Real" } GT_Contact(in1 := #HMI_AnalogValveControl.rManualSP, in2 := #crMaxSetPoint)
      { S7_GenerateENO := "TRUE" } Move(in := #crMaxSetPoint, out1 => #HMI_AnalogValveControl.rManualSP)
      wire#w1
      Coil( #bTemp )
   END_RUNG
   RUNG wire#powerrail
      { S7_Templates := "SrcType := Real" } LT_Contact(in1 := #HMI_AnalogValveControl.rManualSP, in2 := #crMinSetPoint)
      { S7_GenerateENO := "TRUE" } Move(in := #crMinSetPoint, out1 => #HMI_AnalogValveControl.rManualSP)
   END_RUNG wire#w1
   RUNG wire#powerrail
      { S7_Templates := "SrcType := Real" } GT_Contact(in1 := #HMI_AnalogValveControl.rAutoSP, in2 := #crMaxSetPoint)
      { S7_GenerateENO := "TRUE" } Move(in := #crMaxSetPoint, out1 => #HMI_AnalogValveControl.rAutoSP)
   END_RUNG wire#w1
   RUNG wire#powerrail
      { S7_Templates := "SrcType := Real" } LT_Contact(in1 := #HMI_AnalogValveControl.rAutoSP, in2 := #crMinSetPoint)
      { S7_GenerateENO := "TRUE" } Move(in := #crMinSetPoint, out1 => #HMI_AnalogValveControl.rAutoSP)
   END_RUNG wire#w1
   // the same network as SCL:
   // ENO of a box is taken as its EN; it also drops when the box reports an error
   #_w1 := #HMI_AnalogValveControl.rManualSP > #crMaxSetPoint;
   IF #_w1 THEN #HMI_AnalogValveControl.rManualSP := #crMaxSetPoint; END_IF;
   #_w2 := #HMI_AnalogValveControl.rManualSP < #crMinSetPoint;
   IF #_w2 THEN #HMI_AnalogValveControl.rManualSP := #crMinSetPoint; END_IF;
   #_w3 := #HMI_AnalogValveControl.rAutoSP > #crMaxSetPoint;
   IF #_w3 THEN #HMI_AnalogValveControl.rAutoSP := #crMaxSetPoint; END_IF;
   #_w4 := #HMI_AnalogValveControl.rAutoSP < #crMinSetPoint;
   IF #_w4 THEN #HMI_AnalogValveControl.rAutoSP := #crMinSetPoint; END_IF;
   #bTemp := #_w1 OR #_w2 OR #_w3 OR #_w4;
END_REGION

REGION Network 6: Reset Errors
   RUNG wire#powerrail
      Contact( #bInResetError )
      wire#w1
      Contact( #HMI_AnalogValveControl.bPBEN_ResetError )
      Coil( #bReset )
      R_Coil( #ERROR_AnalogValve.InvalidFeedback )
   END_RUNG
   RUNG wire#powerrail
      Contact( #bPB_ResetError )
   END_RUNG wire#w1
   // the same network as SCL:
   #bReset := (#bInResetError OR #bPB_ResetError) AND #HMI_AnalogValveControl.bPBEN_ResetError;
   IF #bReset THEN #ERROR_AnalogValve.InvalidFeedback := FALSE; END_IF;
END_REGION

REGION Network 7: Set mode override if neccesary
   RUNG wire#powerrail
      { S7_Templates := "SrcType := Int" } NE_Contact(in1 := #iInMode, in2 := "Modes.Independent")
      { S7_GenerateENO := "TRUE" } Move(in := #iInMode, out1 => #HMI_AnalogValveControl.iMode)
   END_RUNG
   // the same network as SCL:
   IF #iInMode <> "Modes.Independent" THEN #HMI_AnalogValveControl.iMode := #iInMode; END_IF;
END_REGION

REGION Network 8: Enable the reset error pushbutton if there is an error
   RUNG wire#powerrail
      Contact( #HMI_AnalogValveControl.bError )
      Coil( #HMI_AnalogValveControl.bPBEN_ResetError )
   END_RUNG
   // the same network as SCL:
   #HMI_AnalogValveControl.bPBEN_ResetError := #HMI_AnalogValveControl.bError;
END_REGION

REGION Network 9: Set actual value based on mode